(* Logix 5000 project; controller PLC_MCC1300_75F1 vendor 1 type 14 code 166 rev 32.11; software revision 32.04; part 24 of 83 *)
(* tags used below, declared in another part *)
   GP_M316A : GP_Rotator;
   M302SpeedUp : MAC_SpeedUp;
   M310B : MAC_Conveyor;
   M315A : MAC_Conveyor;
   M315B : MAC_Conveyor;
   M316 : MAC_Conveyor;
   M316_ALM : MAC_Conveyor_ALM;
   M316_Data : UDT_Convoy_SL;
   M316_HMR : MAC_Conveyor_HMR;
   M316_HMW : MAC_Conveyor_HMW;
   M316_M1_DR : AXIS_CIP_DRIVE;
   M316_M1_DR_IN_MAJ : MOTION_INSTRUCTION;
   M316_M1_DR_IN_MAR : MOTION_INSTRUCTION;
   M316_M1_DR_IN_MAS : MOTION_INSTRUCTION;
   M316_M1_DR_IN_MRP : MOTION_INSTRUCTION;
   M316_M1_DR_MAFR : MOTION_INSTRUCTION;
   M316_M1_DR_MDR : MOTION_INSTRUCTION;
   M316_M1_DR_MSF : MOTION_INSTRUCTION;
   M316_M1_DR_MSO : MOTION_INSTRUCTION;
   M316_M1_DR_OUT_MAJ : MOTION_INSTRUCTION;
   M316_M1_DR_OUT_MAM : MOTION_INSTRUCTION;
   M316_M1_DR_OUT_MAR : MOTION_INSTRUCTION;
   M316_M1_DR_OUT_MAS : MOTION_INSTRUCTION;
   M316_M1_DR_OUT_MCD : MOTION_INSTRUCTION;
   M316_M1_DR_OUT_MRP : MOTION_INSTRUCTION;
   M316_SpaceConv_Utilities : SpaceConv_Utilities;
   M316A : MAC_Rotator;
   M316A_HMR : MAC_Rotator_HMR;
   M316A_HMW : MAC_Rotator_HMW;
   M316A_M1_DR : AXIS_CIP_DRIVE;
   M316A_M1_DR_IN_MAM : MOTION_INSTRUCTION;
   M316A_M1_DR_IN_MAS : MOTION_INSTRUCTION;
   M316A_M1_DR_MAFR : MOTION_INSTRUCTION;
   M316A_M1_DR_MAH : MOTION_INSTRUCTION;
   M316A_M1_DR_MSF : MOTION_INSTRUCTION;
   M316A_M1_DR_MSO : MOTION_INSTRUCTION;
   M316A_M1_DR_OUT_MAJ : MOTION_INSTRUCTION;
   M316A_M1_DR_OUT_MAM : MOTION_INSTRUCTION;
   M316A_M1_DR_OUT_MAS : MOTION_INSTRUCTION;
   M316A_MAM_IP_TOFF : TIMER;
   M317 : MAC_Conveyor_Single;
   TMP_d : DINT;
   TMP_dDirection : DINT;
   TMP_r : REAL;
   TMP_rAcc : REAL;
   TMP_rDec : REAL;
   TMP_rSpeed : REAL;
   TMP_rTarget : REAL;
   TMP_rTarget_M1 : REAL;
   TMP_xForwardCommadnForCleaningZone : BOOL;
   TMP_xPositioning : BOOL;
   TMP_xPositioning_M1 : BOOL;
   TMP_xPowerSaving : BOOL;
   TMP_xReverse : BOOL;
   TMP_xReverse_M1 : BOOL;
   TMP_xRun : BOOL;
   TMP_xRun_M1 : BOOL;
   xAlwaysOFF : BOOL;
   xDebugOFF : BOOL;
   Z300_Conveyor : UDT_StandConv[29];
   Z300_Conveyor_Conf : UDT_Conveyor_Config[29];
   Z300_Conveyor_HMW : MAC_Conveyor_ZC_HMW[29];
   Z300_Conveyor_IN_MOTION : MAC_Conveyor_ZC_IN_MOTION[29];
   Z301_HMR : MAC_Zone_ML_HMR;
   Z401 : MAC_Zone;
   Z402 : MAC_Zone;
   Z402_HMW : MAC_Zone_HMW;
(* CommandLogic, continued *)

ROUTINE M315M3_Conveyor_Output   (* ladder *)
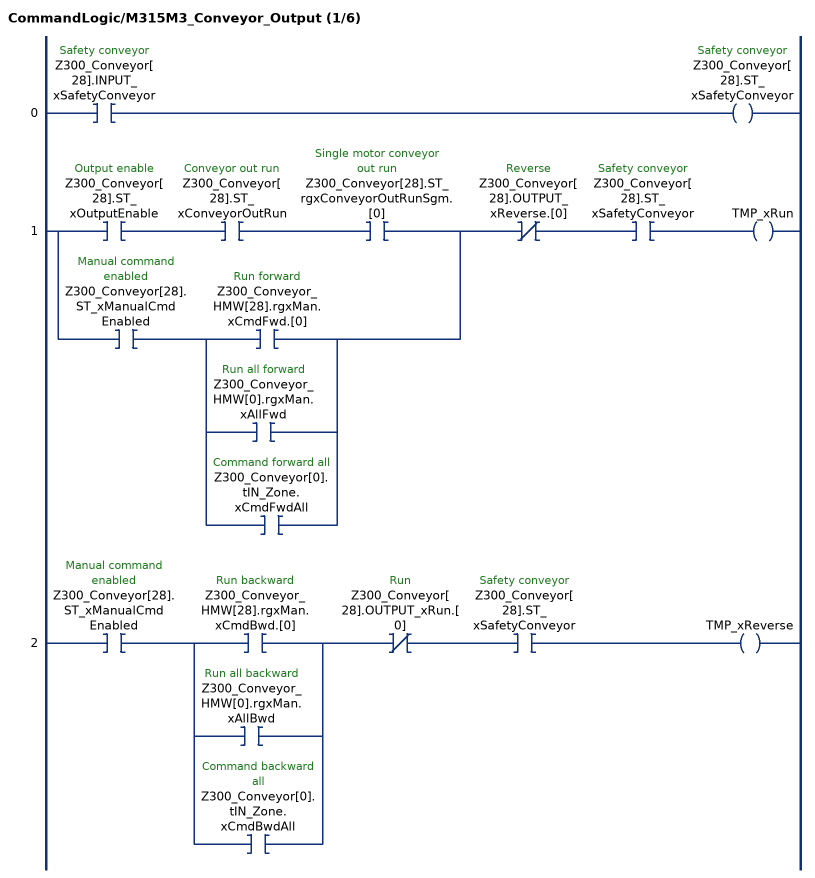
   0: XIC(Z300_Conveyor[28].INPUT_xSafetyConveyor)OTE(Z300_Conveyor[28].ST_xSafetyConveyor);
   1: [XIC(Z300_Conveyor[28].ST_xOutputEnable) XIC(Z300_Conveyor[28].ST_xConveyorOutRun) XIC(Z300_Conveyor[28].ST_rgxConveyorOutRunSgm.[0]) ,XIC(Z300_Conveyor[28].ST_xManualCmdEnabled) [XIC(Z300_Conveyor_HMW[28].rgxMan.xCmdFwd.[0]) ,XIC(Z300_Conveyor_HMW[0].rgxMan.xAllFwd) ,XIC(Z300_Conveyor[0].tIN_Zone.xCmdFwdAll) ] ]XIO(Z300_Conveyor[28].OUTPUT_xReverse.[0])XIC(Z300_Conveyor[28].ST_xSafetyConveyor)OTE(TMP_xRun);
   2: XIC(Z300_Conveyor[28].ST_xManualCmdEnabled)[XIC(Z300_Conveyor_HMW[28].rgxMan.xCmdBwd.[0]) ,XIC(Z300_Conveyor_HMW[0].rgxMan.xAllBwd) ,XIC(Z300_Conveyor[0].tIN_Zone.xCmdBwdAll) ]XIO(Z300_Conveyor[28].OUTPUT_xRun.[0])XIC(Z300_Conveyor[28].ST_xSafetyConveyor)OTE(TMP_xReverse);
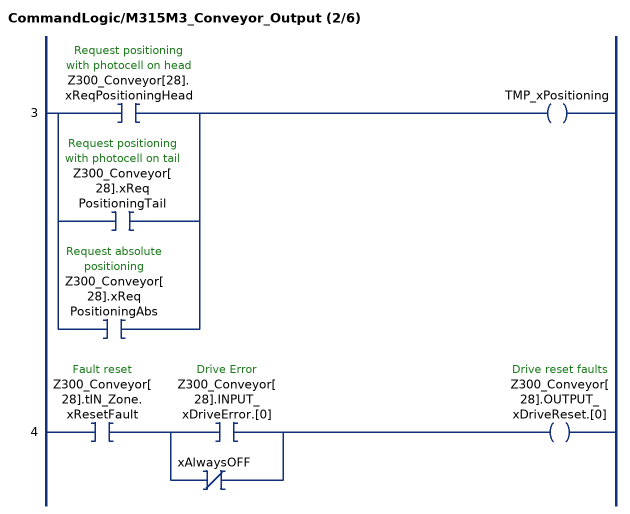
   3: [XIC(Z300_Conveyor[28].xReqPositioningHead) ,XIC(Z300_Conveyor[28].xReqPositioningTail) ,XIC(Z300_Conveyor[28].xReqPositioningAbs) ]OTE(TMP_xPositioning);
   4: XIC(Z300_Conveyor[28].tIN_Zone.xResetFault)[XIC(Z300_Conveyor[28].INPUT_xDriveError.[0]) ,XIO(xAlwaysOFF) ]OTE(Z300_Conveyor[28].OUTPUT_xDriveReset.[0]);
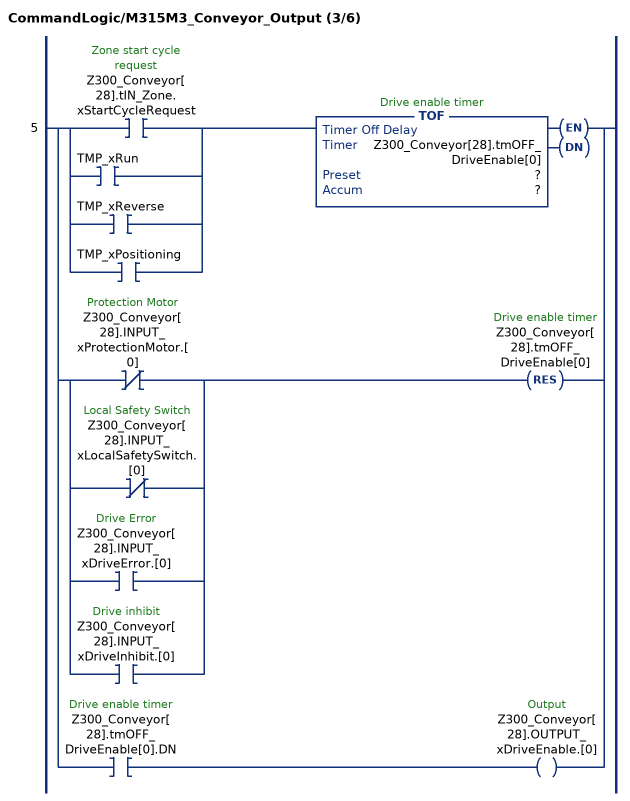
   5: [[XIC(Z300_Conveyor[28].tIN_Zone.xStartCycleRequest) ,XIC(TMP_xRun) ,XIC(TMP_xReverse) ,XIC(TMP_xPositioning) ] TOF(Z300_Conveyor[28].tmOFF_DriveEnable[0],?,?) ,[XIO(Z300_Conveyor[28].INPUT_xProtectionMotor.[0]) ,XIO(Z300_Conveyor[28].INPUT_xLocalSafetySwitch.[0]) ,XIC(Z300_Conveyor[28].INPUT_xDriveError.[0]) ,XIC(Z300_Conveyor[28].INPUT_xDriveInhibit.[0]) ] RES(Z300_Conveyor[28].tmOFF_DriveEnable[0]) ,XIC(Z300_Conveyor[28].tmOFF_DriveEnable[0].DN) OTE(Z300_Conveyor[28].OUTPUT_xDriveEnable.[0]) ];
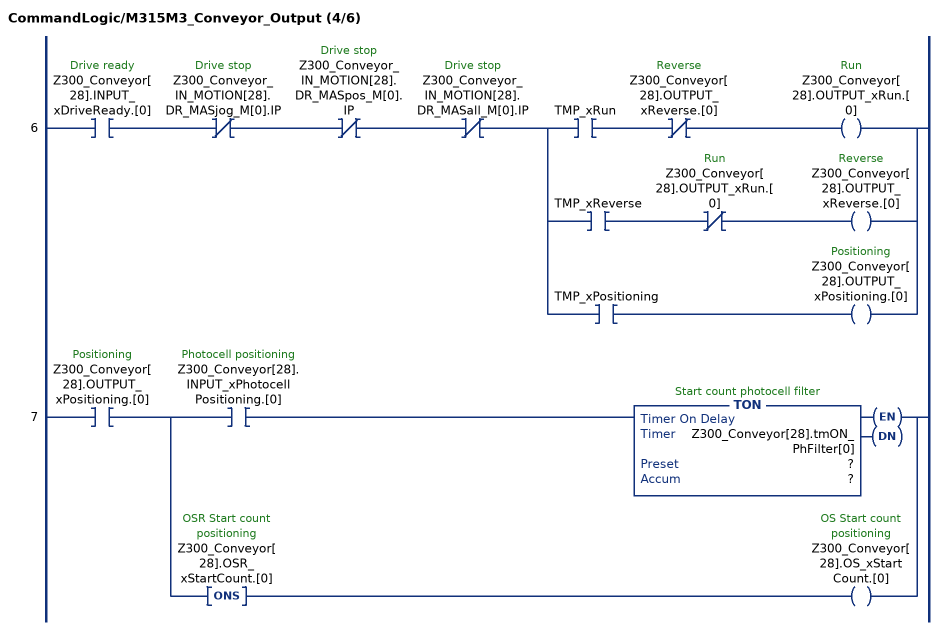
   6: XIC(Z300_Conveyor[28].INPUT_xDriveReady.[0])XIO(Z300_Conveyor_IN_MOTION[28].DR_MASjog_M[0].IP)XIO(Z300_Conveyor_IN_MOTION[28].DR_MASpos_M[0].IP)XIO(Z300_Conveyor_IN_MOTION[28].DR_MASall_M[0].IP)[XIC(TMP_xRun) XIO(Z300_Conveyor[28].OUTPUT_xReverse.[0]) OTE(Z300_Conveyor[28].OUTPUT_xRun.[0]) ,XIC(TMP_xReverse) XIO(Z300_Conveyor[28].OUTPUT_xRun.[0]) OTE(Z300_Conveyor[28].OUTPUT_xReverse.[0]) ,XIC(TMP_xPositioning) OTE(Z300_Conveyor[28].OUTPUT_xPositioning.[0]) ];
   7: XIC(Z300_Conveyor[28].OUTPUT_xPositioning.[0])[XIC(Z300_Conveyor[28].INPUT_xPhotocellPositioning.[0]) TON(Z300_Conveyor[28].tmON_PhFilter[0],?,?) ,ONS(Z300_Conveyor[28].OSR_xStartCount.[0]) OTE(Z300_Conveyor[28].OS_xStartCount.[0]) ];
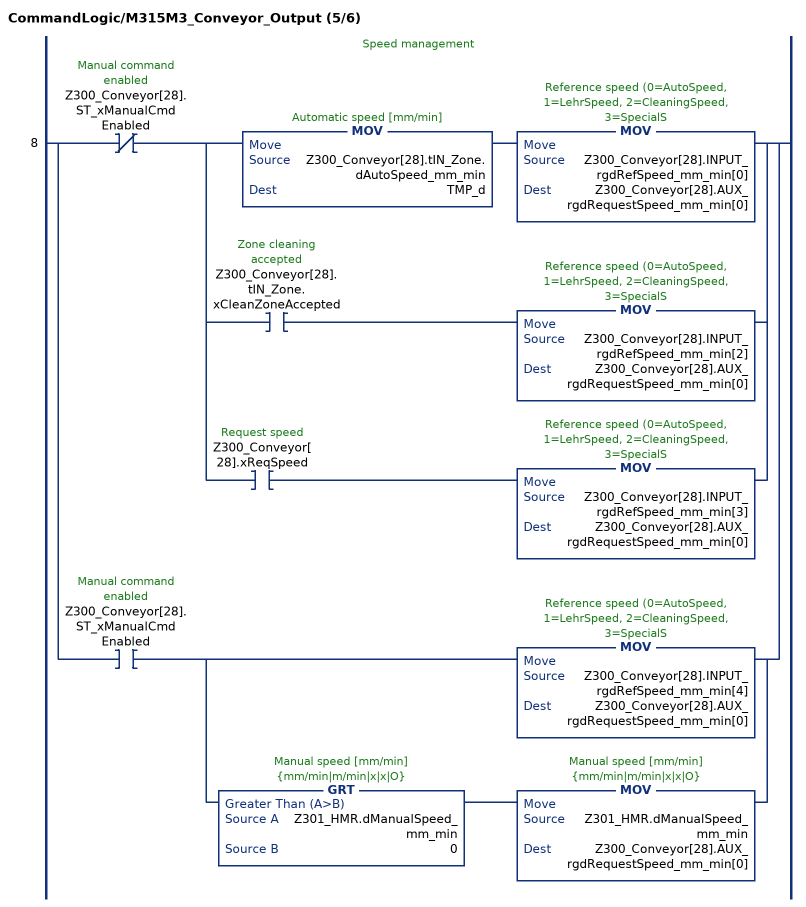
   // Speed management
   8: [XIO(Z300_Conveyor[28].ST_xManualCmdEnabled) [MOV(Z300_Conveyor[28].tIN_Zone.dAutoSpeed_mm_min,TMP_d) MOV(Z300_Conveyor[28].INPUT_rgdRefSpeed_mm_min[0],Z300_Conveyor[28].AUX_rgdRequestSpeed_mm_min[0]) ,XIC(Z300_Conveyor[28].tIN_Zone.xCleanZoneAccepted) MOV(Z300_Conveyor[28].INPUT_rgdRefSpeed_mm_min[2],Z300_Conveyor[28].AUX_rgdRequestSpeed_mm_min[0]) ,XIC(Z300_Conveyor[28].xReqSpeed) MOV(Z300_Conveyor[28].INPUT_rgdRefSpeed_mm_min[3],Z300_Conveyor[28].AUX_rgdRequestSpeed_mm_min[0]) ] ,XIC(Z300_Conveyor[28].ST_xManualCmdEnabled) [MOV(Z300_Conveyor[28].INPUT_rgdRefSpeed_mm_min[4],Z300_Conveyor[28].AUX_rgdRequestSpeed_mm_min[0]) ,GRT(Z301_HMR.dManualSpeed_mm_min,0) MOV(Z301_HMR.dManualSpeed_mm_min,Z300_Conveyor[28].AUX_rgdRequestSpeed_mm_min[0]) ] ];
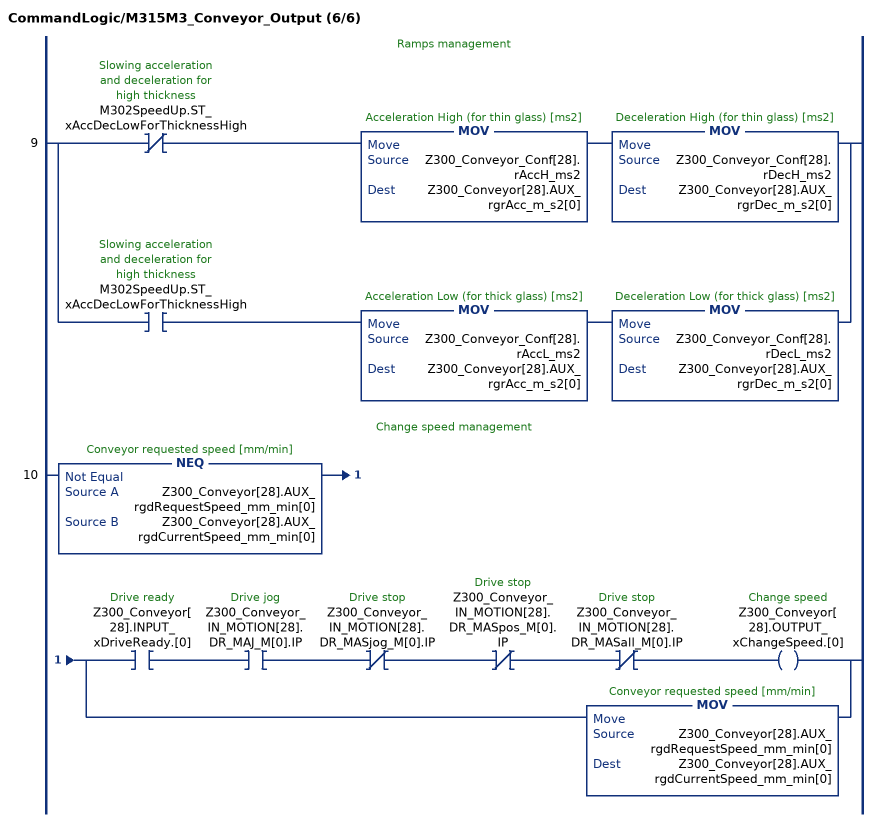
   // Ramps management
   9: [XIO(M302SpeedUp.ST_xAccDecLowForThicknessHigh) MOV(Z300_Conveyor_Conf[28].rAccH_ms2,Z300_Conveyor[28].AUX_rgrAcc_m_s2[0]) MOV(Z300_Conveyor_Conf[28].rDecH_ms2,Z300_Conveyor[28].AUX_rgrDec_m_s2[0]) ,XIC(M302SpeedUp.ST_xAccDecLowForThicknessHigh) MOV(Z300_Conveyor_Conf[28].rAccL_ms2,Z300_Conveyor[28].AUX_rgrAcc_m_s2[0]) MOV(Z300_Conveyor_Conf[28].rDecL_ms2,Z300_Conveyor[28].AUX_rgrDec_m_s2[0]) ];
   // Change speed management
   10: NEQ(Z300_Conveyor[28].AUX_rgdRequestSpeed_mm_min[0],Z300_Conveyor[28].AUX_rgdCurrentSpeed_mm_min[0])[XIC(Z300_Conveyor[28].INPUT_xDriveReady.[0]) XIC(Z300_Conveyor_IN_MOTION[28].DR_MAJ_M[0].IP) XIO(Z300_Conveyor_IN_MOTION[28].DR_MASjog_M[0].IP) XIO(Z300_Conveyor_IN_MOTION[28].DR_MASpos_M[0].IP) XIO(Z300_Conveyor_IN_MOTION[28].DR_MASall_M[0].IP) OTE(Z300_Conveyor[28].OUTPUT_xChangeSpeed.[0]) ,MOV(Z300_Conveyor[28].AUX_rgdRequestSpeed_mm_min[0],Z300_Conveyor[28].AUX_rgdCurrentSpeed_mm_min[0]) ];
END_ROUTINE

ROUTINE M316_Output   (* ladder *)
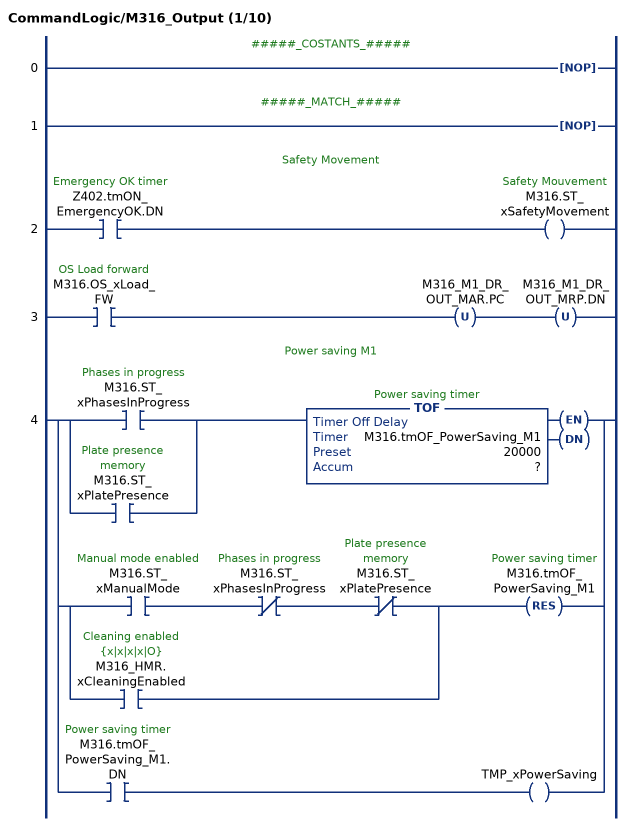
   // #####_COSTANTS_#####
   0: NOP();
   // #####_MATCH_#####
   1: NOP();
   // Safety Movement
   2: XIC(Z402.tmON_EmergencyOK.DN)OTE(M316.ST_xSafetyMovement);
   3: XIC(M316.OS_xLoad_FW)OTU(M316_M1_DR_OUT_MAR.PC)OTU(M316_M1_DR_OUT_MRP.DN);
   // Power saving M1
   4: [[XIC(M316.ST_xPhasesInProgress) ,XIC(M316.ST_xPlatePresence) ] TOF(M316.tmOF_PowerSaving_M1,?,?) ,[XIC(M316.ST_xManualMode) XIO(M316.ST_xPhasesInProgress) XIO(M316.ST_xPlatePresence) ,XIC(M316_HMR.xCleaningEnabled) ] RES(M316.tmOF_PowerSaving_M1) ,XIC(M316.tmOF_PowerSaving_M1.DN) OTE(TMP_xPowerSaving) ];
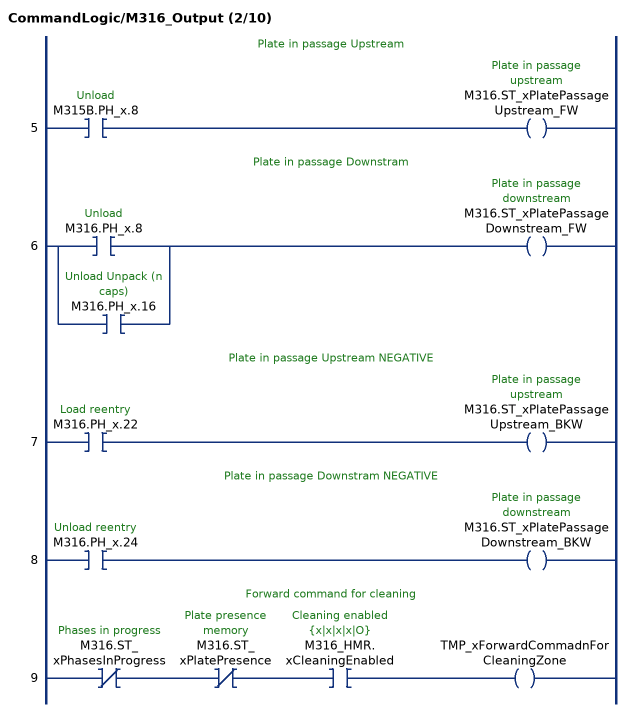
   // Plate in passage Upstream
   5: XIC(M315B.PH_x.8)OTE(M316.ST_xPlatePassageUpstream_FW);
   // Plate in passage Downstram
   6: [XIC(M316.PH_x.8) ,XIC(M316.PH_x.16) ]OTE(M316.ST_xPlatePassageDownstream_FW);
   // Plate in passage Upstream NEGATIVE
   7: XIC(M316.PH_x.22)OTE(M316.ST_xPlatePassageUpstream_BKW);
   // Plate in passage Downstram NEGATIVE
   8: XIC(M316.PH_x.24)OTE(M316.ST_xPlatePassageDownstream_BKW);
   // Forward command for cleaning
   9: XIO(M316.ST_xPhasesInProgress)XIO(M316.ST_xPlatePresence)XIC(M316_HMR.xCleaningEnabled)OTE(TMP_xForwardCommadnForCleaningZone);
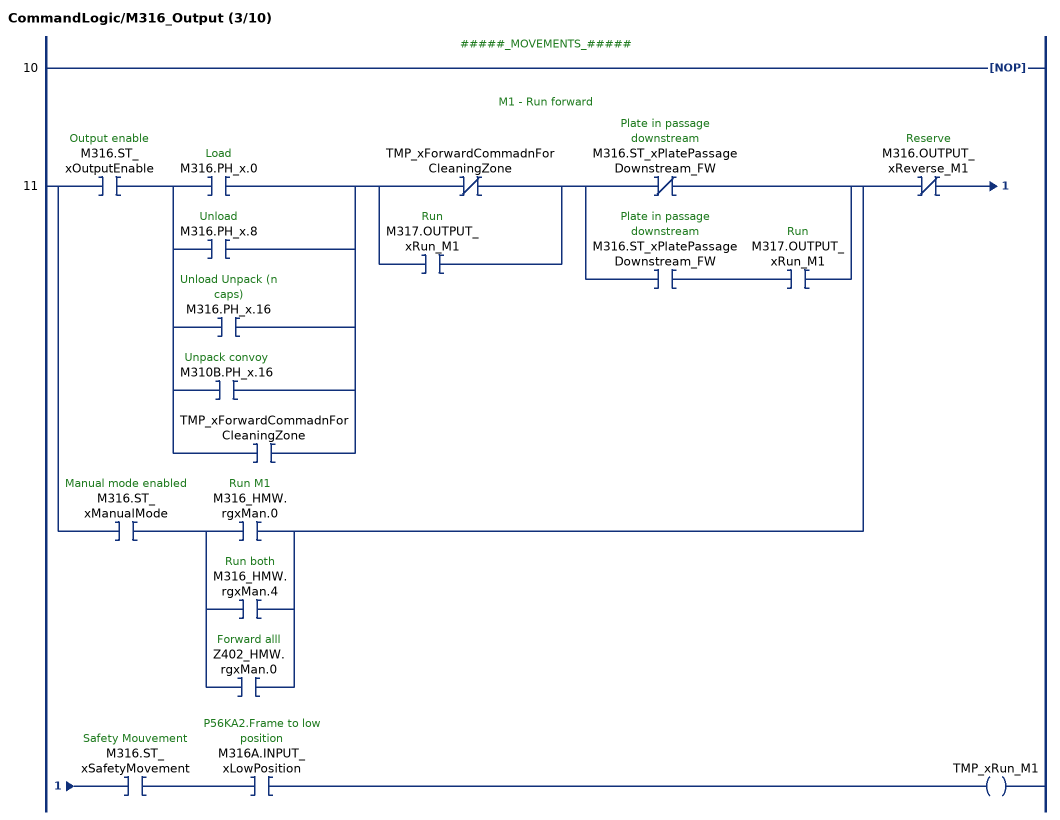
   // #####_MOVEMENTS_#####
   10: NOP();
   // M1 - Run forward
   11: [XIC(M316.ST_xOutputEnable) [XIC(M316.PH_x.0) ,XIC(M316.PH_x.8) ,XIC(M316.PH_x.16) ,XIC(M310B.PH_x.16) ,XIC(TMP_xForwardCommadnForCleaningZone) ] [XIO(TMP_xForwardCommadnForCleaningZone) ,XIC(M317.OUTPUT_xRun_M1) ] [XIO(M316.ST_xPlatePassageDownstream_FW) ,XIC(M316.ST_xPlatePassageDownstream_FW) XIC(M317.OUTPUT_xRun_M1) ] ,XIC(M316.ST_xManualMode) [XIC(M316_HMW.rgxMan.0) ,XIC(M316_HMW.rgxMan.4) ,XIC(Z402_HMW.rgxMan.0) ] ]XIO(M316.OUTPUT_xReverse_M1)XIC(M316.ST_xSafetyMovement)XIC(M316A.INPUT_xLowPosition)OTE(TMP_xRun_M1);
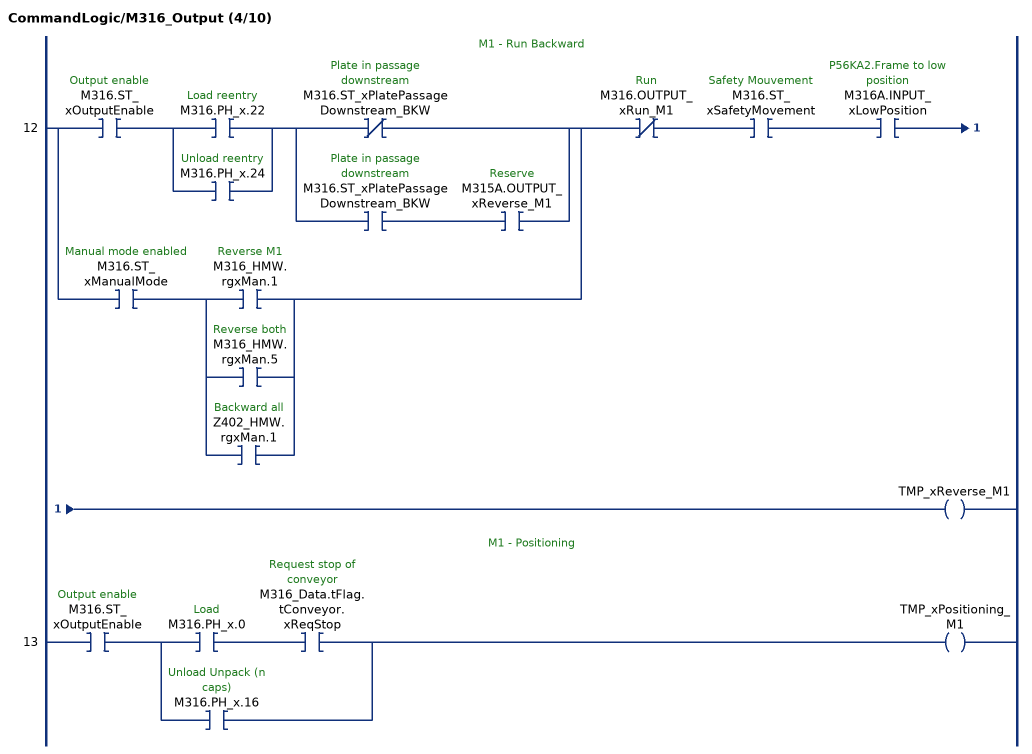
   // M1 - Run Backward
   12: [XIC(M316.ST_xOutputEnable) [XIC(M316.PH_x.22) ,XIC(M316.PH_x.24) ] [XIO(M316.ST_xPlatePassageDownstream_BKW) ,XIC(M316.ST_xPlatePassageDownstream_BKW) XIC(M315A.OUTPUT_xReverse_M1) ] ,XIC(M316.ST_xManualMode) [XIC(M316_HMW.rgxMan.1) ,XIC(M316_HMW.rgxMan.5) ,XIC(Z402_HMW.rgxMan.1) ] ]XIO(M316.OUTPUT_xRun_M1)XIC(M316.ST_xSafetyMovement)XIC(M316A.INPUT_xLowPosition)OTE(TMP_xReverse_M1);
   // M1 - Positioning
   13: XIC(M316.ST_xOutputEnable)[XIC(M316.PH_x.0) XIC(M316_Data.tFlag.tConveyor.xReqStop) ,XIC(M316.PH_x.16) ]OTE(TMP_xPositioning_M1);
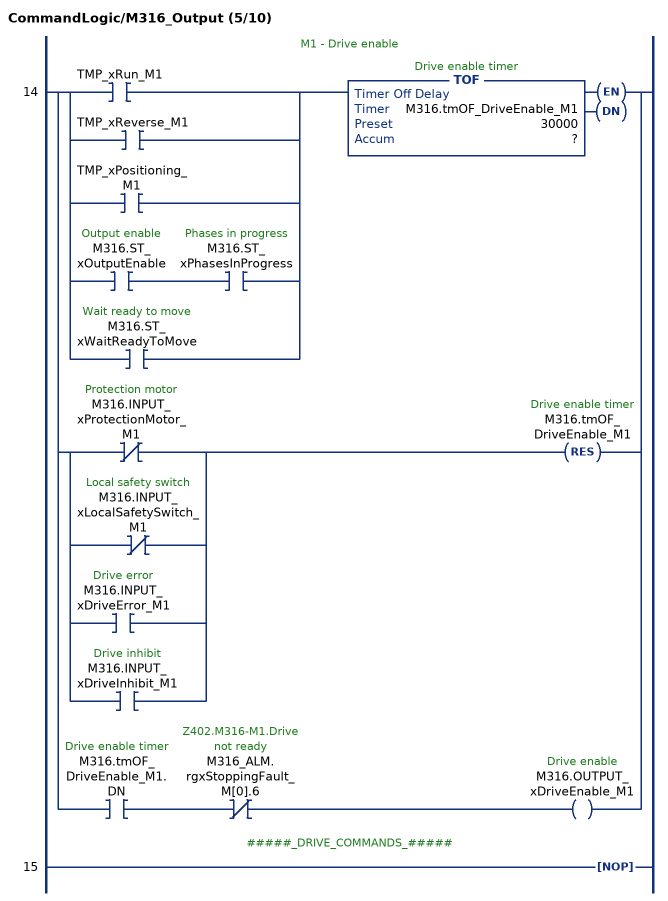
   // M1 - Drive enable
   14: [[XIC(TMP_xRun_M1) ,XIC(TMP_xReverse_M1) ,XIC(TMP_xPositioning_M1) ,XIC(M316.ST_xOutputEnable) XIC(M316.ST_xPhasesInProgress) ,XIC(M316.ST_xWaitReadyToMove) ] TOF(M316.tmOF_DriveEnable_M1,?,?) ,[XIO(M316.INPUT_xProtectionMotor_M1) ,XIO(M316.INPUT_xLocalSafetySwitch_M1) ,XIC(M316.INPUT_xDriveError_M1) ,XIC(M316.INPUT_xDriveInhibit_M1) ] RES(M316.tmOF_DriveEnable_M1) ,XIC(M316.tmOF_DriveEnable_M1.DN) XIO(M316_ALM.rgxStoppingFault_M[0].6) OTE(M316.OUTPUT_xDriveEnable_M1) ];
   // #####_DRIVE_COMMANDS_#####
   15: NOP();
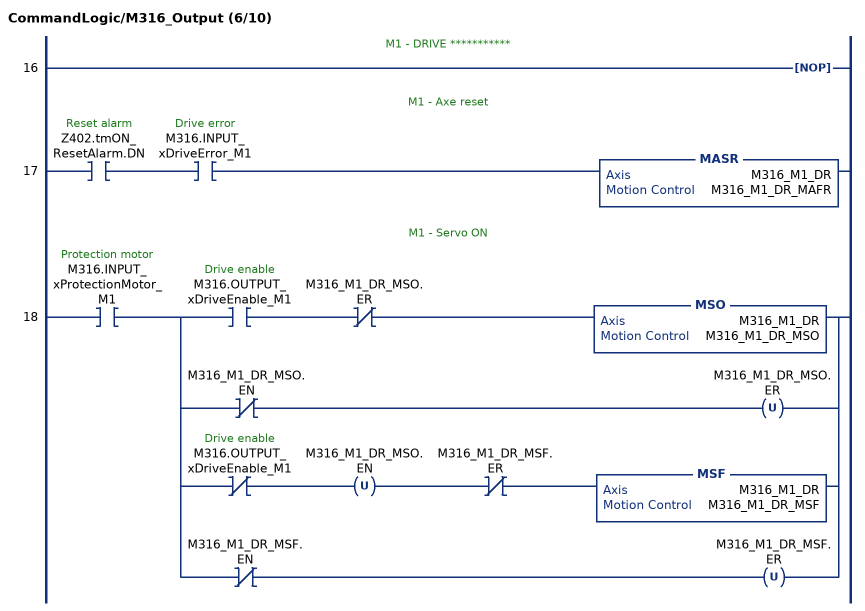
   // M1 - DRIVE ***********
   16: NOP();
   // M1 - Axe reset
   17: XIC(Z402.tmON_ResetAlarm.DN)XIC(M316.INPUT_xDriveError_M1)MASR(M316_M1_DR,M316_M1_DR_MAFR);
   // M1 - Servo ON
   18: XIC(M316.INPUT_xProtectionMotor_M1)[XIC(M316.OUTPUT_xDriveEnable_M1) XIO(M316_M1_DR_MSO.ER) MSO(M316_M1_DR,M316_M1_DR_MSO) ,XIO(M316_M1_DR_MSO.EN) OTU(M316_M1_DR_MSO.ER) ,XIO(M316.OUTPUT_xDriveEnable_M1) OTU(M316_M1_DR_MSO.EN) XIO(M316_M1_DR_MSF.ER) MSF(M316_M1_DR,M316_M1_DR_MSF) ,XIO(M316_M1_DR_MSF.EN) OTU(M316_M1_DR_MSF.ER) ];